(* Logix 5000 project; controller FV vendor 1 type 14 code 217 rev 31.11; software revision 31.00; part 11 of 63 *)
(* tags used below, declared in another part *)
   CWD : CHECKWORD_FLAGS;
   FR_B230 : INT[255];   // FLOW_BITS Flow Meter Bits
   FR_B240 : INT[255];   // DEBOUNCE Debounce Flags
   FR_B246 : INT[255];   // V_REVERSE Flags for reversing contol action
   FR_CFG1_P : PlantItem;   // CFG1_P
   FR_CFG2_P : PlantItem;   // CFG2_P
   FR_data_file_value_to_move : DINT;
   FR_FILT_PR_PX : PlantItem;   // FILT_PR_PX
   FR_FILT_TNK_PX : PlantItem;   // FILT_TNK_PX
   FR_FILT_TNLN_PX : PlantItem;   // FILT_TNLN_PX
   FR_FRV1_AV01 : PlantItem;   // FRV1_AV01
   FR_FV26_AV01 : PlantItem;   // FV26_AV01
   FR_FV26_AV04 : PlantItem;   // FV26_AV04
   FR_FV26_AV05 : PlantItem;   // FV26_AV05
   FR_FV26_AV06 : PlantItem;   // FV26_AV06
   FR_FV26_AV07 : PlantItem;   // FV26_AV07
   FR_FV26_VA01 : PlantItem;   // FV26_VA01
   FR_FV27_AV04 : PlantItem;   // FV27_AV04
   FR_FV28_AV04 : PlantItem;   // FV28_AV04
   FR_FV29_AV04 : PlantItem;   // FV29_AV04
   FR_FV30_AV04 : PlantItem;   // FV30_AV04
   FR_FV31_AV04 : PlantItem;   // FV31_AV04
   FR_FVR1_P01 : PlantItem;   // FVR1_P01
   FR_N10 : INT[265];   // FV_AGING Comms to FV Aging PL C
   FR_N100 : INT[265];   // FV FILLING
   FR_N110 : INT[265];   // GREEN BEER Green Beer Main
   FR_N120 : INT[265];   // YEAST CROP Yeast Cropping Main
   FR_N13 : INT[265];   // MV_ROUTE Comms to MV Routing PLC
   FR_N130 : INT[265];   // FILTRATE Filtrate Return
   FR_N14 : INT[265];   // MVFV CIP Comms to MVFV CIP Un it PLC
   FR_N160 : INT[265];   // VESSEL Vessel Working Direc tory
   FR_N200 : INT[265];   // ANALOG_IN Analog Inputs
   FR_N255 : INT[265];   // CHECKWORDS
   FR_N26 : INT[265];   // FV26
   FR_N7 : INT[265];   // INTEGER
   FR_N99 : INT[265];   // COMMENT Comment Lines
   FR_PANELESTOP : PlantItem;   // PANELESTOP
   FR_PARAF : PlantItem;   // PARAF
   FR_PILZ : PlantItem;   // PILZ
   FR_T131 : TIMER[255];   // FILTRATE
   FR_T144 : TIMER[255];   // CIP
   FR_T4 : TIMER[255];   // TIMER
   FR_VB1_AV08 : PlantItem;   // VB1_AV08
   FR_VB1_AV09 : PlantItem;   // VB1_AV09
   FR_VB4_AV01 : PlantItem;   // VB4_AV01
   FR_VB4_AV07 : PlantItem;   // VB4_AV07
   FR_VB4_AV13 : PlantItem;   // VB4_AV13
   FR_VB4_AV19 : PlantItem;   // VB4_AV19
   FR_VB4_AV21 : PlantItem;   // VB4_AV21
   FR_VB4_AV23 : PlantItem;   // VB4_AV23
(* FR_Common, continued *)

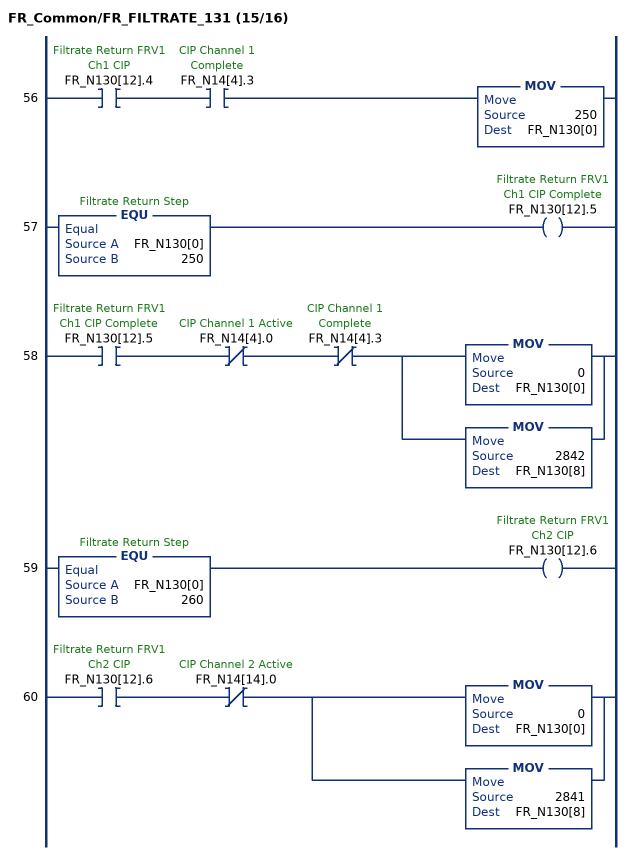
   [picture p136: FR_Common/FR_FILTRATE_131 rungs 56-60]
   56: XIC(FR_N130[12].4)XIC(FR_N14[4].3)MOV(250,FR_N130[0]);
   57: EQU(FR_N130[0],250)OTE(FR_N130[12].5);
   58: XIC(FR_N130[12].5)XIO(FR_N14[4].0)XIO(FR_N14[4].3)[MOV(0,FR_N130[0]) ,MOV(2842,FR_N130[8]) ];
   59: EQU(FR_N130[0],260)OTE(FR_N130[12].6);
   60: XIC(FR_N130[12].6)XIO(FR_N14[14].0)[MOV(0,FR_N130[0]) ,MOV(2841,FR_N130[8]) ];
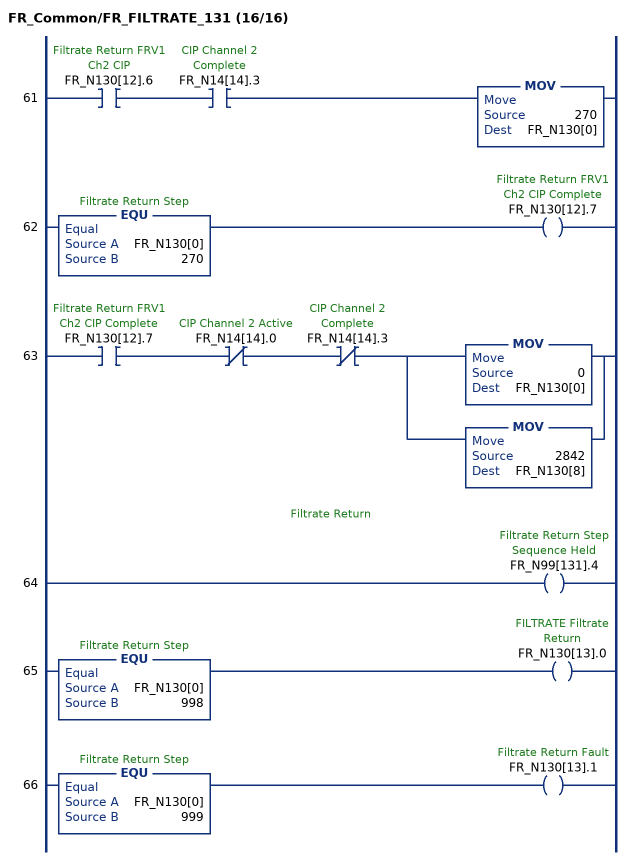
   61: XIC(FR_N130[12].6)XIC(FR_N14[14].3)MOV(270,FR_N130[0]);
   62: EQU(FR_N130[0],270)OTE(FR_N130[12].7);
   63: XIC(FR_N130[12].7)XIO(FR_N14[14].0)XIO(FR_N14[14].3)[MOV(0,FR_N130[0]) ,MOV(2842,FR_N130[8]) ];
   // Filtrate Return
   64: OTE(FR_N99[131].4);
   65: EQU(FR_N130[0],998)OTE(FR_N130[13].0);
   66: EQU(FR_N130[0],999)OTE(FR_N130[13].1);
END_ROUTINE

ROUTINE FR_FILTRATE_O_132   (* ladder *)
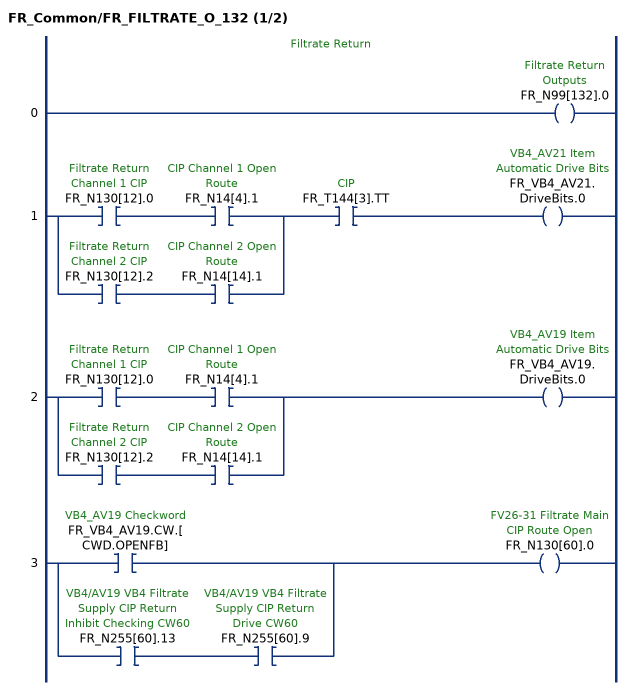
   // Filtrate Return
   0: OTE(FR_N99[132].0);
   1: [XIC(FR_N130[12].0) XIC(FR_N14[4].1) ,XIC(FR_N130[12].2) XIC(FR_N14[14].1) ]XIC(FR_T144[3].TT)OTE(FR_VB4_AV21.DriveBits.0);
   2: [XIC(FR_N130[12].0) XIC(FR_N14[4].1) ,XIC(FR_N130[12].2) XIC(FR_N14[14].1) ]OTE(FR_VB4_AV19.DriveBits.0);
   3: [XIC(FR_VB4_AV19.CW.[CWD.OPENFB]) ,XIC(FR_N255[60].13) XIC(FR_N255[60].9) ]OTE(FR_N130[60].0);
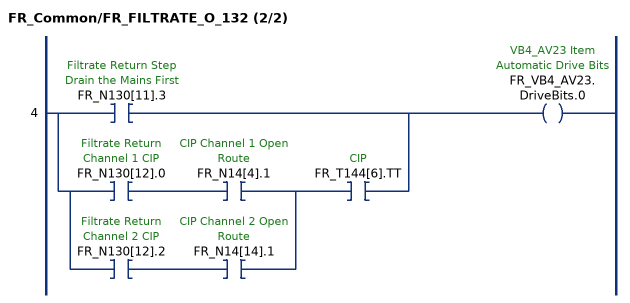
   4: [XIC(FR_N130[11].3) ,[XIC(FR_N130[12].0) XIC(FR_N14[4].1) ,XIC(FR_N130[12].2) XIC(FR_N14[14].1) ] XIC(FR_T144[6].TT) ]OTE(FR_VB4_AV23.DriveBits.0);
END_ROUTINE

ROUTINE FR_FILTRATE_S_130   (* ladder *)
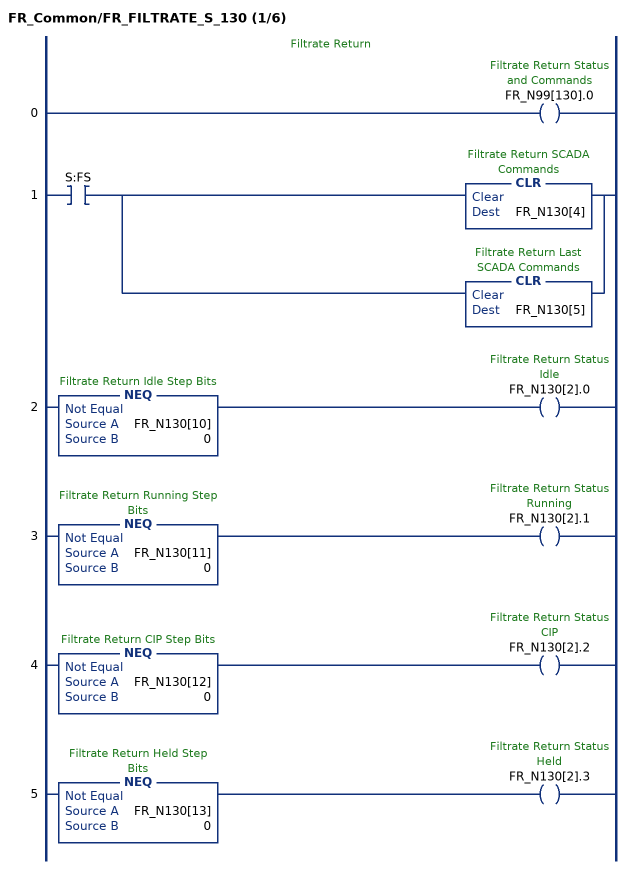
   // Filtrate Return
   0: OTE(FR_N99[130].0);
   1: XIC(S:FS)[CLR(FR_N130[4]) ,CLR(FR_N130[5]) ];
   2: NEQ(FR_N130[10],0)OTE(FR_N130[2].0);
   3: NEQ(FR_N130[11],0)OTE(FR_N130[2].1);
   4: NEQ(FR_N130[12],0)OTE(FR_N130[2].2);
   5: NEQ(FR_N130[13],0)OTE(FR_N130[2].3);
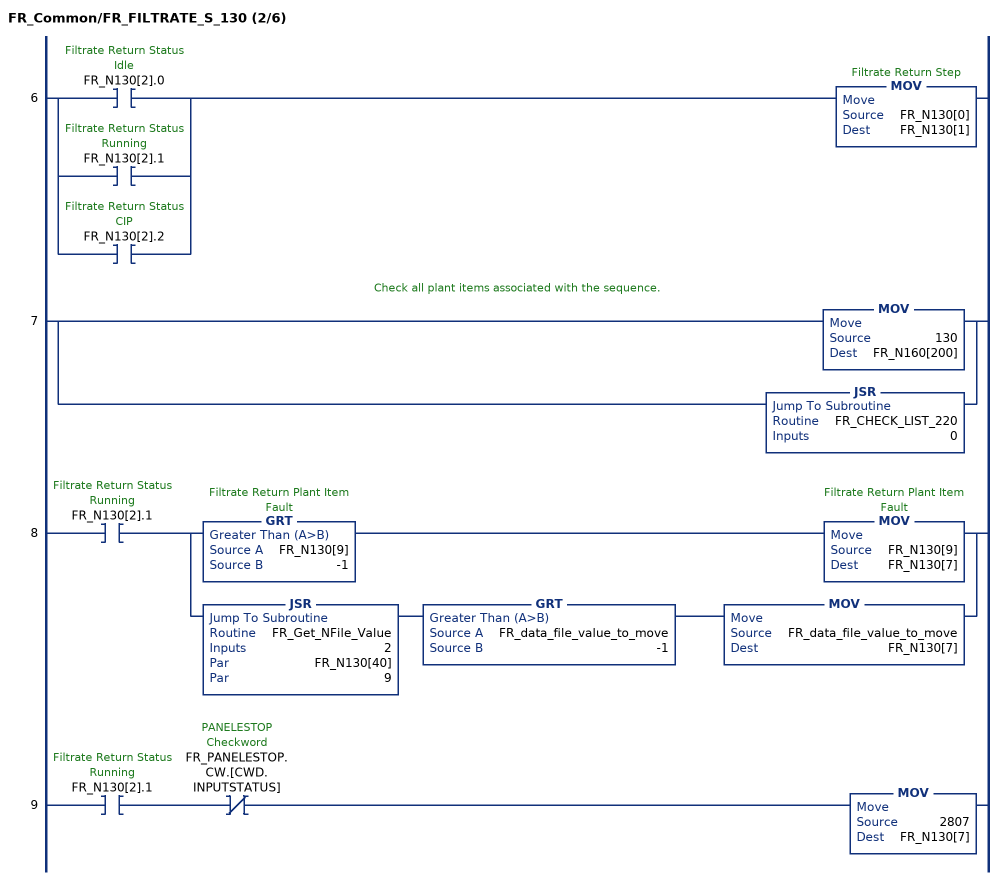
   6: [XIC(FR_N130[2].0) ,XIC(FR_N130[2].1) ,XIC(FR_N130[2].2) ]MOV(FR_N130[0],FR_N130[1]);
   // Check all plant items associated with the sequence.
   7: [MOV(130,FR_N160[200]) ,JSR(FR_CHECK_LIST_220,0) ];
   8: XIC(FR_N130[2].1)[GRT(FR_N130[9],-1) MOV(FR_N130[9],FR_N130[7]) ,JSR(FR_Get_NFile_Value,2,FR_N130[40],9) GRT(FR_data_file_value_to_move,-1) MOV(FR_data_file_value_to_move,FR_N130[7]) ];
   9: XIC(FR_N130[2].1)XIO(FR_PANELESTOP.CW.[CWD.INPUTSTATUS])MOV(2807,FR_N130[7]);
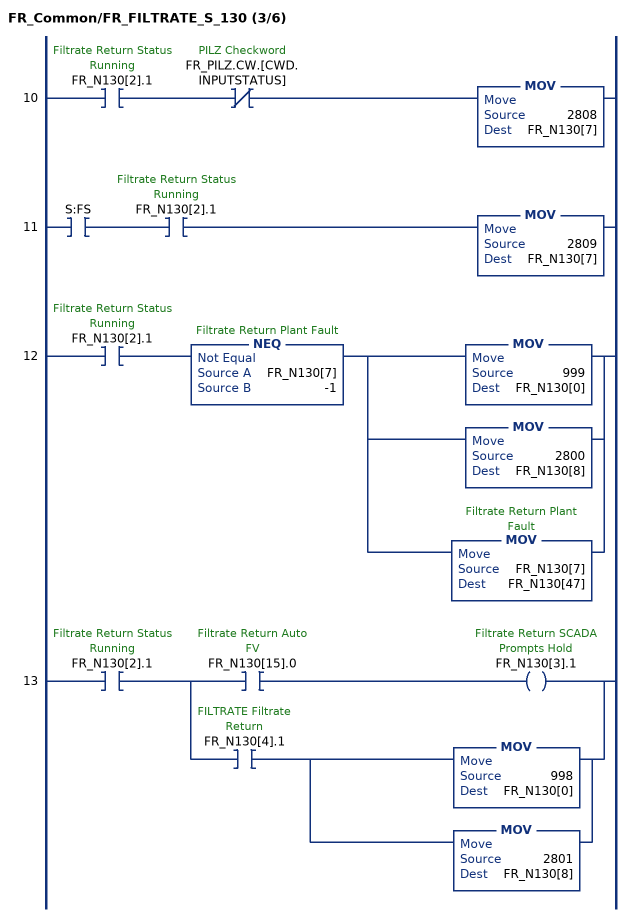
   10: XIC(FR_N130[2].1)XIO(FR_PILZ.CW.[CWD.INPUTSTATUS])MOV(2808,FR_N130[7]);
   11: XIC(S:FS)XIC(FR_N130[2].1)MOV(2809,FR_N130[7]);
   12: XIC(FR_N130[2].1)NEQ(FR_N130[7],-1)[MOV(999,FR_N130[0]) ,MOV(2800,FR_N130[8]) ,MOV(FR_N130[7],FR_N130[47]) ];
   13: XIC(FR_N130[2].1)[XIC(FR_N130[15].0) OTE(FR_N130[3].1) ,XIC(FR_N130[4].1) [MOV(998,FR_N130[0]) ,MOV(2801,FR_N130[8]) ] ];
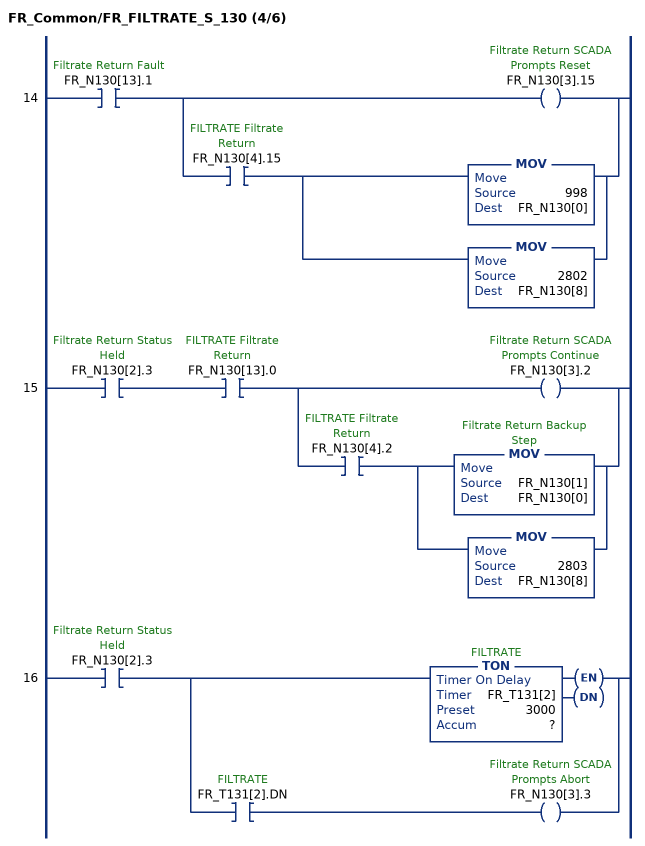
   14: XIC(FR_N130[13].1)[OTE(FR_N130[3].15) ,XIC(FR_N130[4].15) [MOV(998,FR_N130[0]) ,MOV(2802,FR_N130[8]) ] ];
   15: XIC(FR_N130[2].3)XIC(FR_N130[13].0)[OTE(FR_N130[3].2) ,XIC(FR_N130[4].2) [MOV(FR_N130[1],FR_N130[0]) ,MOV(2803,FR_N130[8]) ] ];
   16: XIC(FR_N130[2].3)[TON(FR_T131[2],?,?) ,XIC(FR_T131[2].DN) OTE(FR_N130[3].3) ];
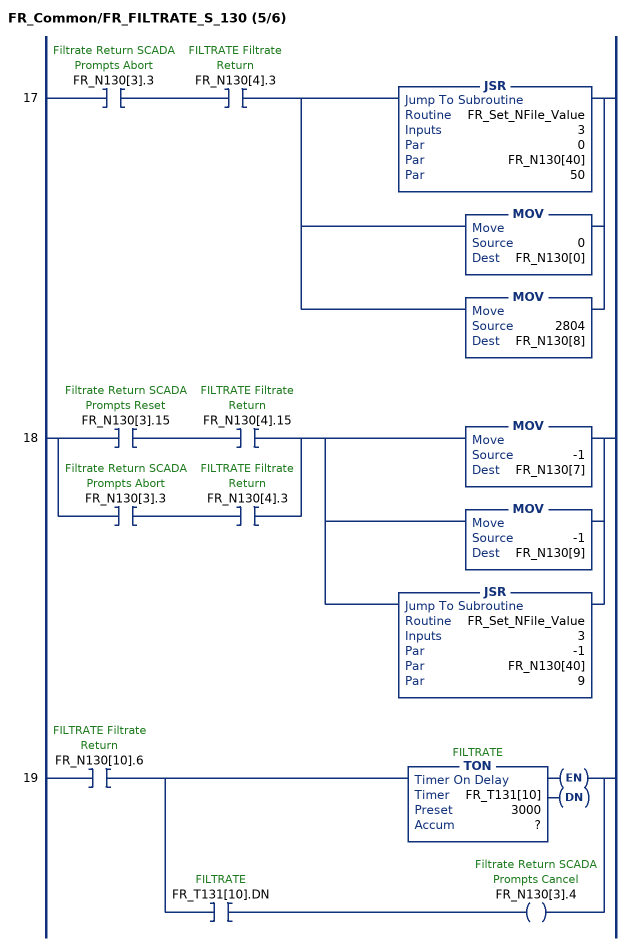
   17: XIC(FR_N130[3].3)XIC(FR_N130[4].3)[JSR(FR_Set_NFile_Value,3,0,FR_N130[40],50) ,MOV(0,FR_N130[0]) ,MOV(2804,FR_N130[8]) ];
   18: [XIC(FR_N130[3].15) XIC(FR_N130[4].15) ,XIC(FR_N130[3].3) XIC(FR_N130[4].3) ][MOV(-1,FR_N130[7]) ,MOV(-1,FR_N130[9]) ,JSR(FR_Set_NFile_Value,3,-1,FR_N130[40],9) ];
   19: XIC(FR_N130[10].6)[TON(FR_T131[10],?,?) ,XIC(FR_T131[10].DN) OTE(FR_N130[3].4) ];
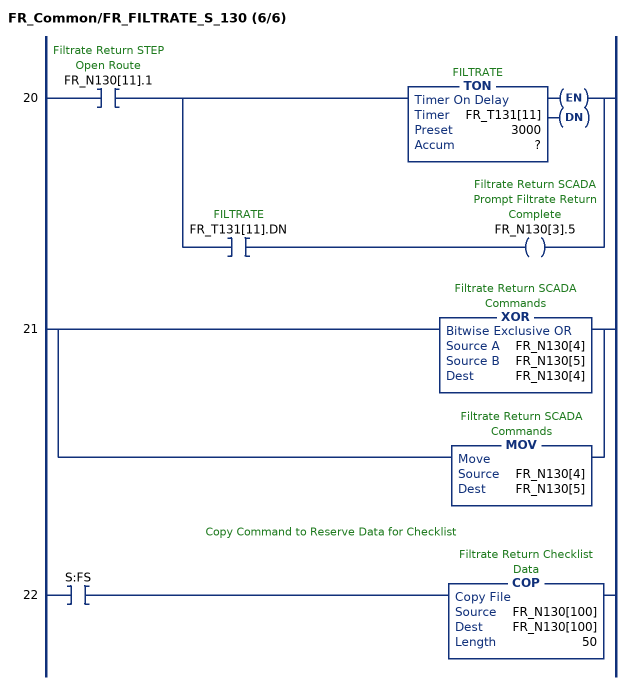
   20: XIC(FR_N130[11].1)[TON(FR_T131[11],?,?) ,XIC(FR_T131[11].DN) OTE(FR_N130[3].5) ];
   21: [XOR(FR_N130[4],FR_N130[5],FR_N130[4]) ,MOV(FR_N130[4],FR_N130[5]) ];
   // Copy Command to Reserve Data for Checklist
   22: XIC(S:FS)COP(FR_N130[100],FR_N130[100],50);
END_ROUTINE

ROUTINE FR_FLOWMETER_230   (* ladder *)
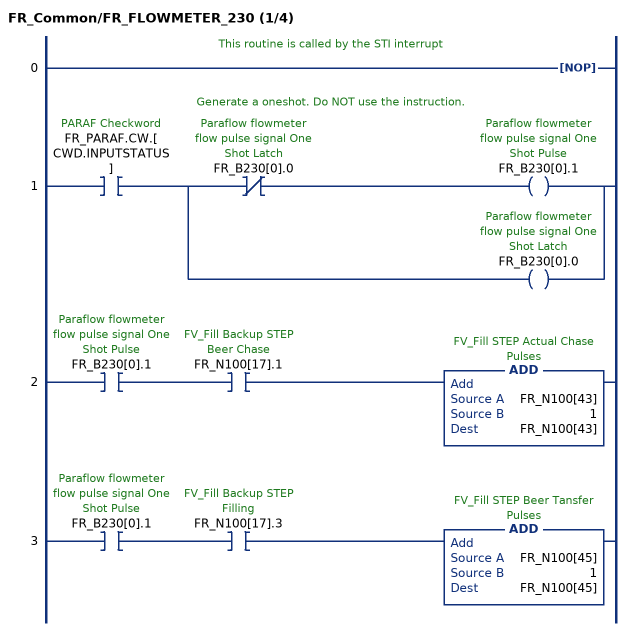
   // This routine is called by the STI interrupt
   0: NOP();
   // Generate a oneshot. Do NOT use the instruction.
   1: XIC(FR_PARAF.CW.[CWD.INPUTSTATUS])[XIO(FR_B230[0].0) OTE(FR_B230[0].1) ,OTE(FR_B230[0].0) ];
   2: XIC(FR_B230[0].1)XIC(FR_N100[17].1)ADD(FR_N100[43],1,FR_N100[43]);
   3: XIC(FR_B230[0].1)XIC(FR_N100[17].3)ADD(FR_N100[45],1,FR_N100[45]);
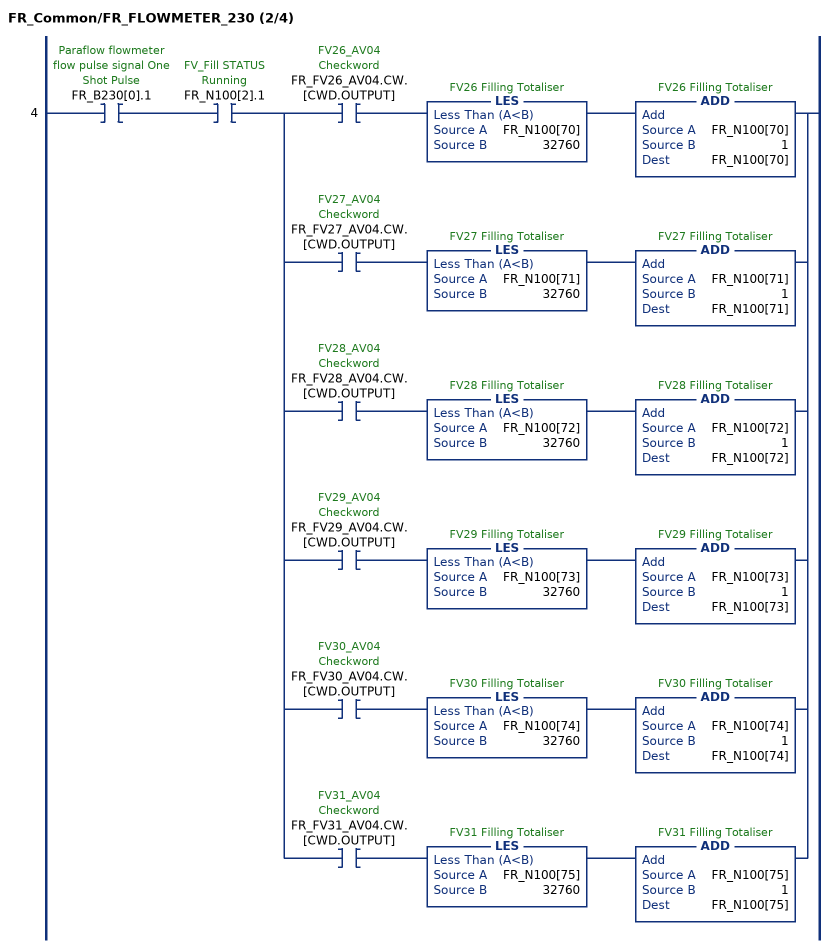
   4: XIC(FR_B230[0].1)XIC(FR_N100[2].1)[XIC(FR_FV26_AV04.CW.[CWD.OUTPUT]) LES(FR_N100[70],32760) ADD(FR_N100[70],1,FR_N100[70]) ,XIC(FR_FV27_AV04.CW.[CWD.OUTPUT]) LES(FR_N100[71],32760) ADD(FR_N100[71],1,FR_N100[71]) ,XIC(FR_FV28_AV04.CW.[CWD.OUTPUT]) LES(FR_N100[72],32760) ADD(FR_N100[72],1,FR_N100[72]) ,XIC(FR_FV29_AV04.CW.[CWD.OUTPUT]) LES(FR_N100[73],32760) ADD(FR_N100[73],1,FR_N100[73]) ,XIC(FR_FV30_AV04.CW.[CWD.OUTPUT]) LES(FR_N100[74],32760) ADD(FR_N100[74],1,FR_N100[74]) ,XIC(FR_FV31_AV04.CW.[CWD.OUTPUT]) LES(FR_N100[75],32760) ADD(FR_N100[75],1,FR_N100[75]) ];
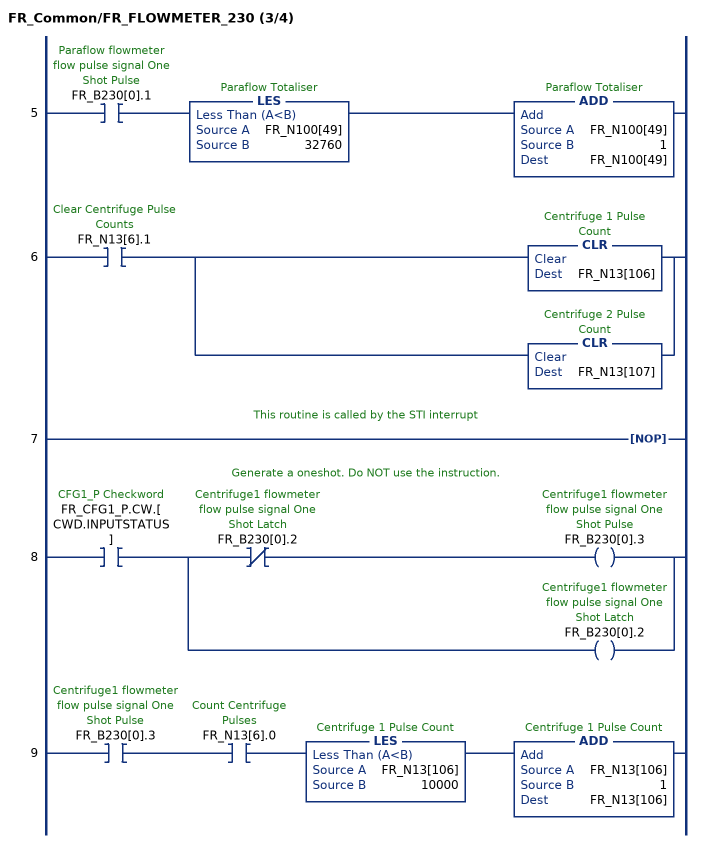
   5: XIC(FR_B230[0].1)LES(FR_N100[49],32760)ADD(FR_N100[49],1,FR_N100[49]);
   6: XIC(FR_N13[6].1)[CLR(FR_N13[106]) ,CLR(FR_N13[107]) ];
   // This routine is called by the STI interrupt
   7: NOP();
   // Generate a oneshot. Do NOT use the instruction.
   8: XIC(FR_CFG1_P.CW.[CWD.INPUTSTATUS])[XIO(FR_B230[0].2) OTE(FR_B230[0].3) ,OTE(FR_B230[0].2) ];
   9: XIC(FR_B230[0].3)XIC(FR_N13[6].0)LES(FR_N13[106],10000)ADD(FR_N13[106],1,FR_N13[106]);
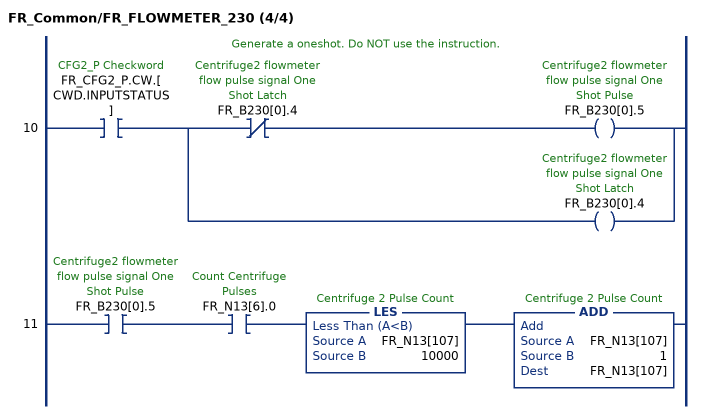
   // Generate a oneshot. Do NOT use the instruction.
   10: XIC(FR_CFG2_P.CW.[CWD.INPUTSTATUS])[XIO(FR_B230[0].4) OTE(FR_B230[0].5) ,OTE(FR_B230[0].4) ];
   11: XIC(FR_B230[0].5)XIC(FR_N13[6].0)LES(FR_N13[107],10000)ADD(FR_N13[107],1,FR_N13[107]);
END_ROUTINE

ROUTINE FR_FRV_133   (* ladder *)
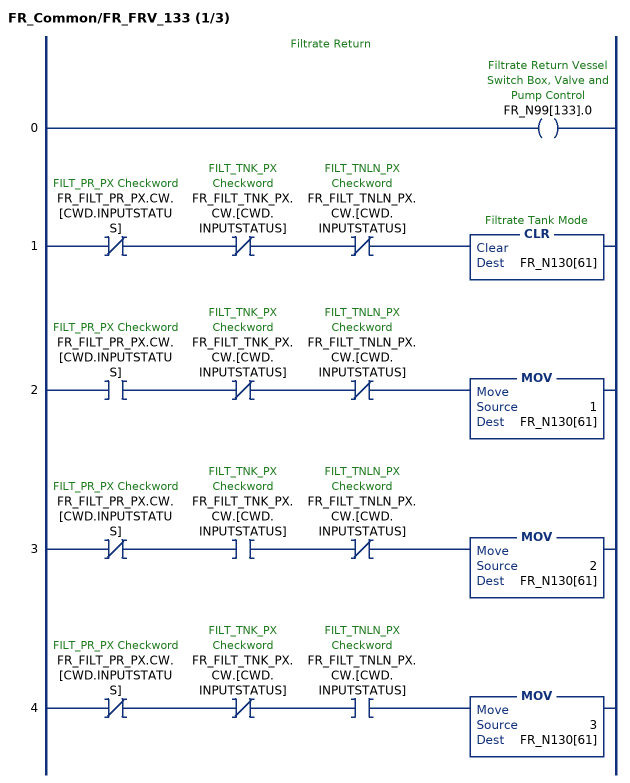
   // Filtrate Return
   0: OTE(FR_N99[133].0);
   1: XIO(FR_FILT_PR_PX.CW.[CWD.INPUTSTATUS])XIO(FR_FILT_TNK_PX.CW.[CWD.INPUTSTATUS])XIO(FR_FILT_TNLN_PX.CW.[CWD.INPUTSTATUS])CLR(FR_N130[61]);
   2: XIC(FR_FILT_PR_PX.CW.[CWD.INPUTSTATUS])XIO(FR_FILT_TNK_PX.CW.[CWD.INPUTSTATUS])XIO(FR_FILT_TNLN_PX.CW.[CWD.INPUTSTATUS])MOV(1,FR_N130[61]);
   3: XIO(FR_FILT_PR_PX.CW.[CWD.INPUTSTATUS])XIC(FR_FILT_TNK_PX.CW.[CWD.INPUTSTATUS])XIO(FR_FILT_TNLN_PX.CW.[CWD.INPUTSTATUS])MOV(2,FR_N130[61]);
   4: XIO(FR_FILT_PR_PX.CW.[CWD.INPUTSTATUS])XIO(FR_FILT_TNK_PX.CW.[CWD.INPUTSTATUS])XIC(FR_FILT_TNLN_PX.CW.[CWD.INPUTSTATUS])MOV(3,FR_N130[61]);
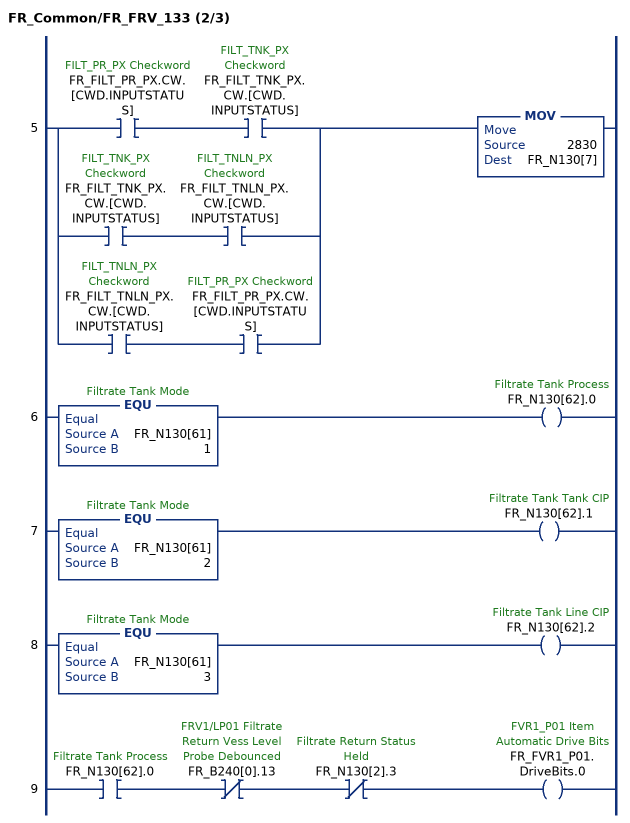
   5: [XIC(FR_FILT_PR_PX.CW.[CWD.INPUTSTATUS]) XIC(FR_FILT_TNK_PX.CW.[CWD.INPUTSTATUS]) ,XIC(FR_FILT_TNK_PX.CW.[CWD.INPUTSTATUS]) XIC(FR_FILT_TNLN_PX.CW.[CWD.INPUTSTATUS]) ,XIC(FR_FILT_TNLN_PX.CW.[CWD.INPUTSTATUS]) XIC(FR_FILT_PR_PX.CW.[CWD.INPUTSTATUS]) ]MOV(2830,FR_N130[7]);
   6: EQU(FR_N130[61],1)OTE(FR_N130[62].0);
   7: EQU(FR_N130[61],2)OTE(FR_N130[62].1);
   8: EQU(FR_N130[61],3)OTE(FR_N130[62].2);
   9: XIC(FR_N130[62].0)XIO(FR_B240[0].13)XIO(FR_N130[2].3)OTE(FR_FVR1_P01.DriveBits.0);
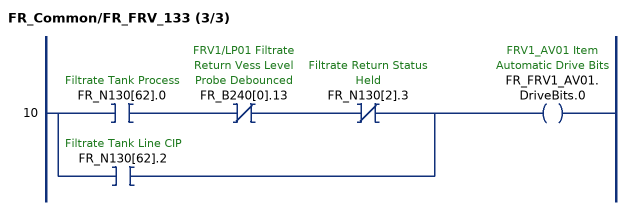
   10: [XIC(FR_N130[62].0) XIO(FR_B240[0].13) XIO(FR_N130[2].3) ,XIC(FR_N130[62].2) ]OTE(FR_FRV1_AV01.DriveBits.0);
END_ROUTINE

ROUTINE FR_FV26_26   (* ladder *)
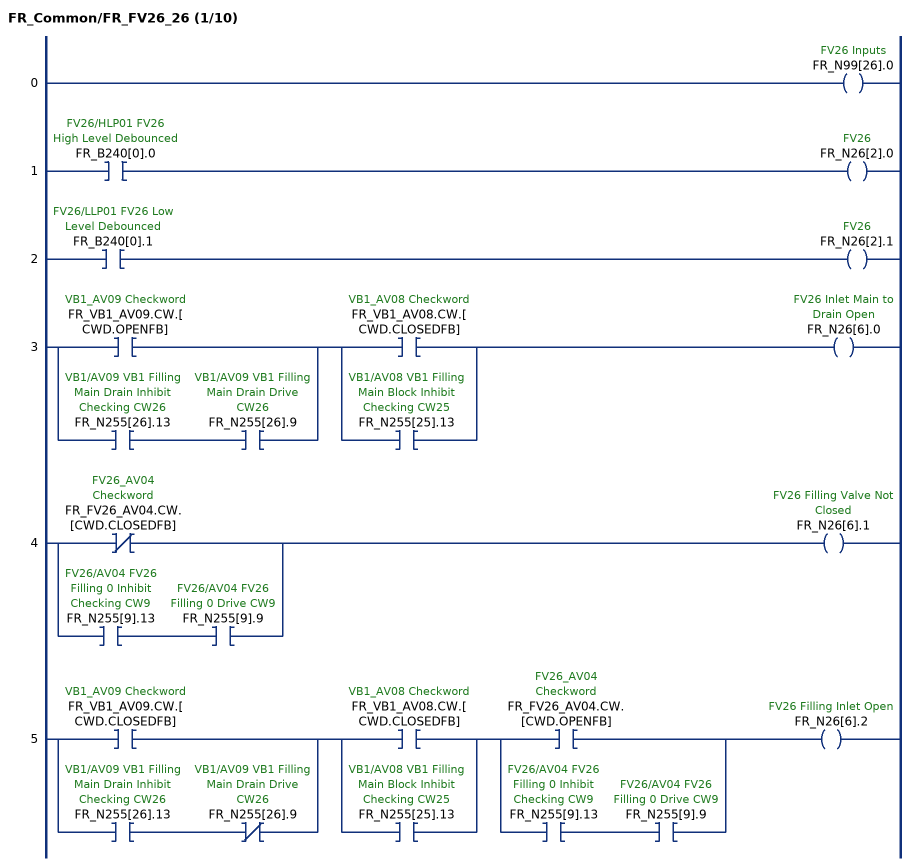
   0: OTE(FR_N99[26].0);
   1: XIC(FR_B240[0].0)OTE(FR_N26[2].0);
   2: XIC(FR_B240[0].1)OTE(FR_N26[2].1);
   3: [XIC(FR_VB1_AV09.CW.[CWD.OPENFB]) ,XIC(FR_N255[26].13) XIC(FR_N255[26].9) ][XIC(FR_VB1_AV08.CW.[CWD.CLOSEDFB]) ,XIC(FR_N255[25].13) ]OTE(FR_N26[6].0);
   4: [XIO(FR_FV26_AV04.CW.[CWD.CLOSEDFB]) ,XIC(FR_N255[9].13) XIC(FR_N255[9].9) ]OTE(FR_N26[6].1);
   5: [XIC(FR_VB1_AV09.CW.[CWD.CLOSEDFB]) ,XIC(FR_N255[26].13) XIO(FR_N255[26].9) ][XIC(FR_VB1_AV08.CW.[CWD.CLOSEDFB]) ,XIC(FR_N255[25].13) ][XIC(FR_FV26_AV04.CW.[CWD.OPENFB]) ,XIC(FR_N255[9].13) XIC(FR_N255[9].9) ]OTE(FR_N26[6].2);
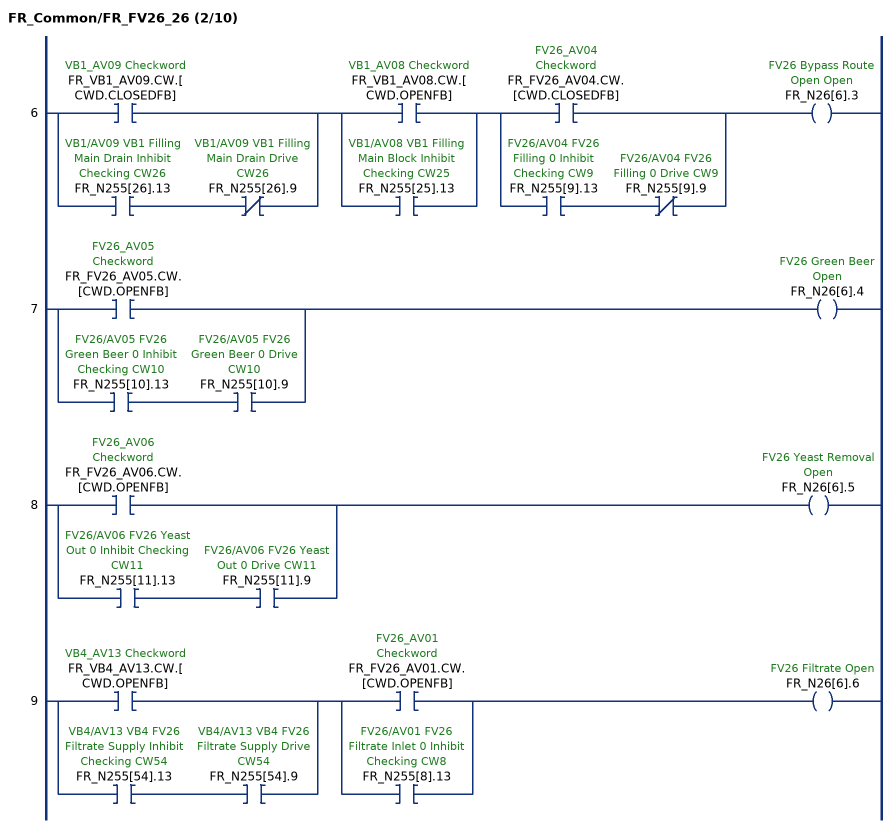
   6: [XIC(FR_VB1_AV09.CW.[CWD.CLOSEDFB]) ,XIC(FR_N255[26].13) XIO(FR_N255[26].9) ][XIC(FR_VB1_AV08.CW.[CWD.OPENFB]) ,XIC(FR_N255[25].13) ][XIC(FR_FV26_AV04.CW.[CWD.CLOSEDFB]) ,XIC(FR_N255[9].13) XIO(FR_N255[9].9) ]OTE(FR_N26[6].3);
   7: [XIC(FR_FV26_AV05.CW.[CWD.OPENFB]) ,XIC(FR_N255[10].13) XIC(FR_N255[10].9) ]OTE(FR_N26[6].4);
   8: [XIC(FR_FV26_AV06.CW.[CWD.OPENFB]) ,XIC(FR_N255[11].13) XIC(FR_N255[11].9) ]OTE(FR_N26[6].5);
   9: [XIC(FR_VB4_AV13.CW.[CWD.OPENFB]) ,XIC(FR_N255[54].13) XIC(FR_N255[54].9) ][XIC(FR_FV26_AV01.CW.[CWD.OPENFB]) ,XIC(FR_N255[8].13) ]OTE(FR_N26[6].6);
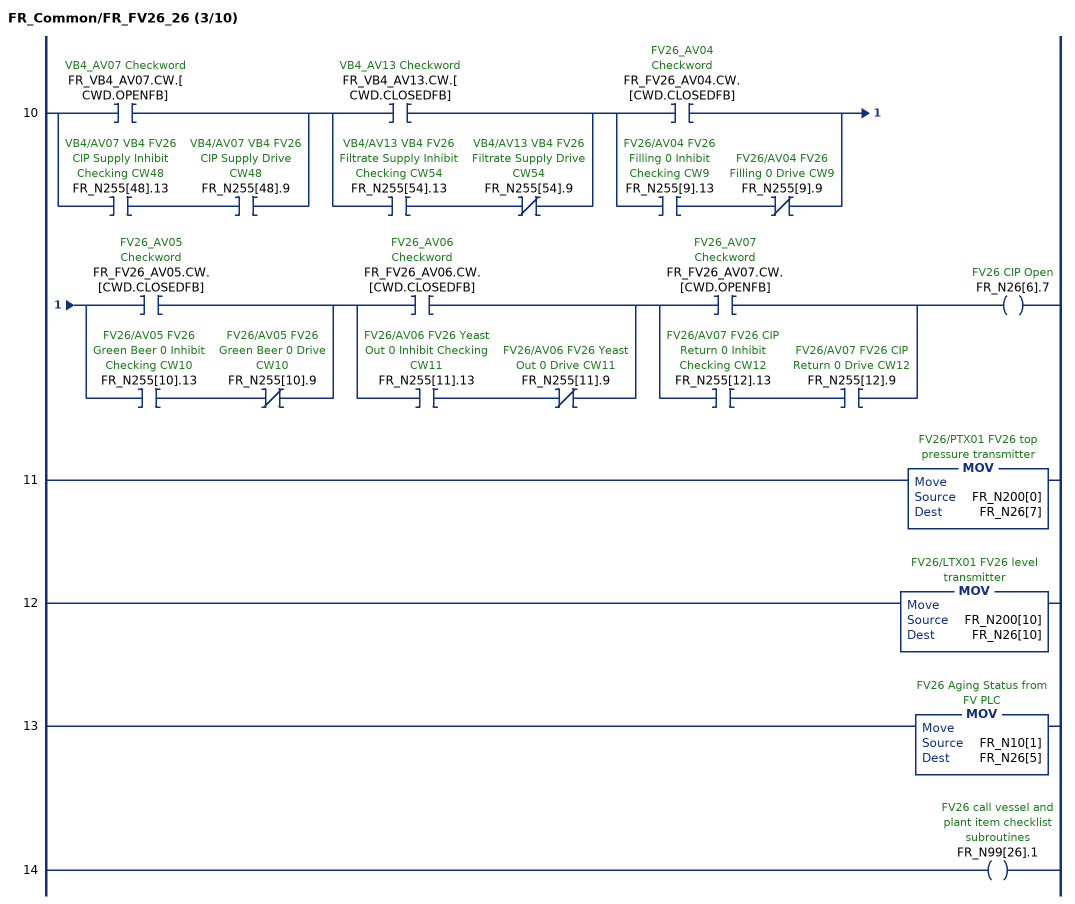
   10: [XIC(FR_VB4_AV07.CW.[CWD.OPENFB]) ,XIC(FR_N255[48].13) XIC(FR_N255[48].9) ][XIC(FR_VB4_AV13.CW.[CWD.CLOSEDFB]) ,XIC(FR_N255[54].13) XIO(FR_N255[54].9) ][XIC(FR_FV26_AV04.CW.[CWD.CLOSEDFB]) ,XIC(FR_N255[9].13) XIO(FR_N255[9].9) ][XIC(FR_FV26_AV05.CW.[CWD.CLOSEDFB]) ,XIC(FR_N255[10].13) XIO(FR_N255[10].9) ][XIC(FR_FV26_AV06.CW.[CWD.CLOSEDFB]) ,XIC(FR_N255[11].13) XIO(FR_N255[11].9) ][XIC(FR_FV26_AV07.CW.[CWD.OPENFB]) ,XIC(FR_N255[12].13) XIC(FR_N255[12].9) ]OTE(FR_N26[6].7);
   11: MOV(FR_N200[0],FR_N26[7]);
   12: MOV(FR_N200[10],FR_N26[10]);
   13: MOV(FR_N10[1],FR_N26[5]);
   14: OTE(FR_N99[26].1);
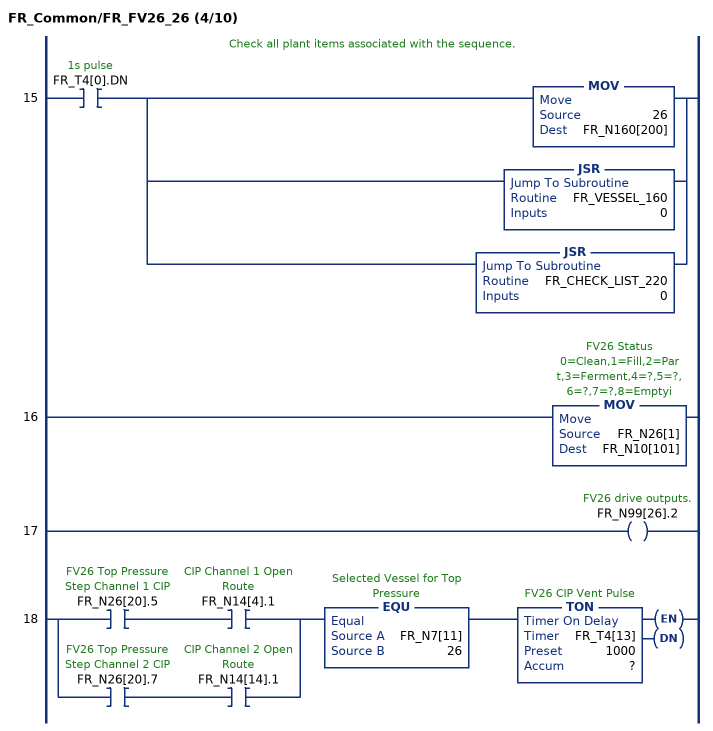
   // Check all plant items associated with the sequence.
   15: XIC(FR_T4[0].DN)[MOV(26,FR_N160[200]) ,JSR(FR_VESSEL_160,0) ,JSR(FR_CHECK_LIST_220,0) ];
   16: MOV(FR_N26[1],FR_N10[101]);
   17: OTE(FR_N99[26].2);
   18: [XIC(FR_N26[20].5) XIC(FR_N14[4].1) ,XIC(FR_N26[20].7) XIC(FR_N14[14].1) ]EQU(FR_N7[11],26)TON(FR_T4[13],?,?);
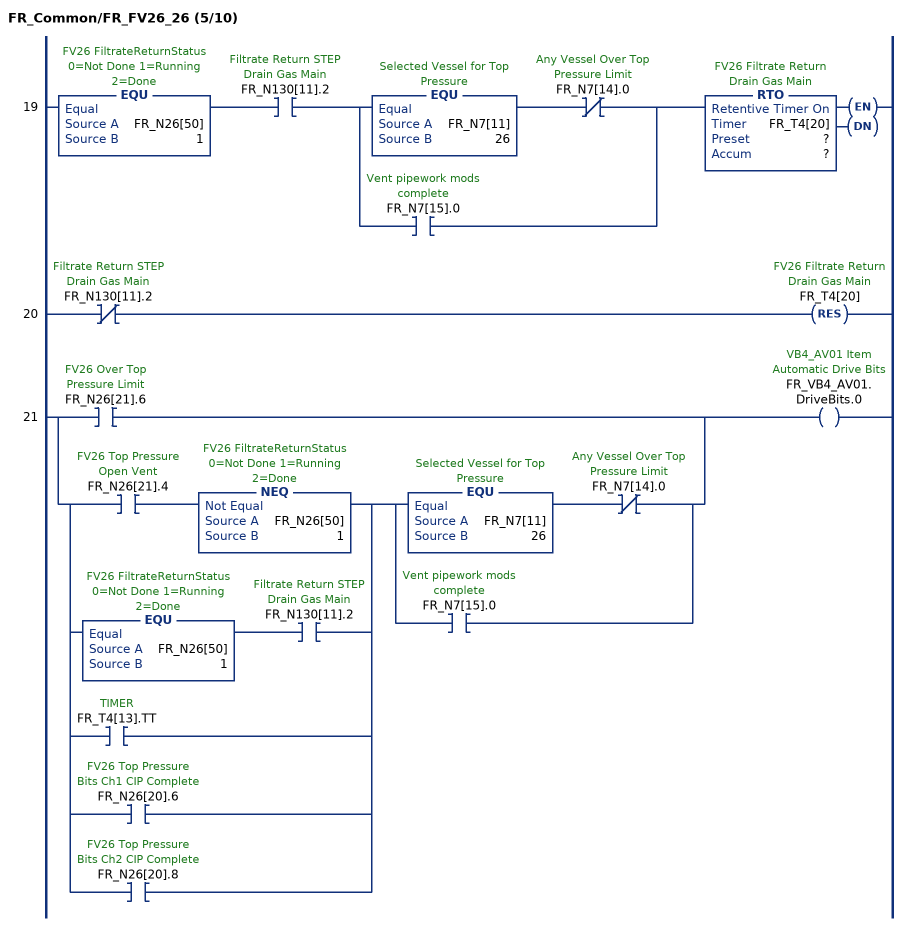
   19: EQU(FR_N26[50],1)XIC(FR_N130[11].2)[EQU(FR_N7[11],26) XIO(FR_N7[14].0) ,XIC(FR_N7[15].0) ]RTO(FR_T4[20],?,?);
   20: XIO(FR_N130[11].2)RES(FR_T4[20]);
   21: [XIC(FR_N26[21].6) ,[XIC(FR_N26[21].4) NEQ(FR_N26[50],1) ,EQU(FR_N26[50],1) XIC(FR_N130[11].2) ,XIC(FR_T4[13].TT) ,[XIC(FR_N26[20].6) ,XIC(FR_N26[20].8) ] ] [EQU(FR_N7[11],26) XIO(FR_N7[14].0) ,XIC(FR_N7[15].0) ] ]OTE(FR_VB4_AV01.DriveBits.0);
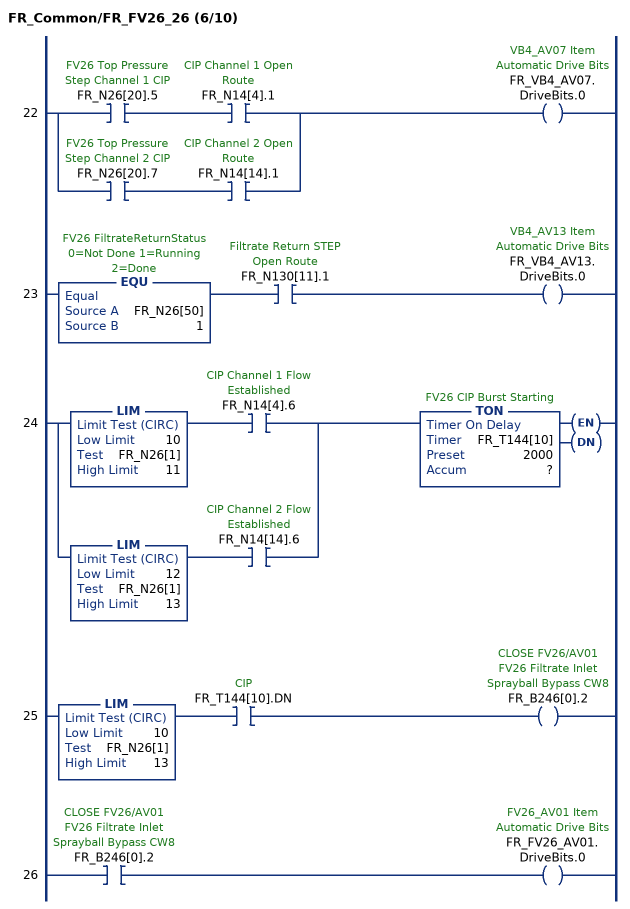
   22: [XIC(FR_N26[20].5) XIC(FR_N14[4].1) ,XIC(FR_N26[20].7) XIC(FR_N14[14].1) ]OTE(FR_VB4_AV07.DriveBits.0);
   23: EQU(FR_N26[50],1)XIC(FR_N130[11].1)OTE(FR_VB4_AV13.DriveBits.0);
   24: [LIM(10,FR_N26[1],11) XIC(FR_N14[4].6) ,LIM(12,FR_N26[1],13) XIC(FR_N14[14].6) ]TON(FR_T144[10],?,?);
   25: LIM(10,FR_N26[1],13)XIC(FR_T144[10].DN)OTE(FR_B246[0].2);
   26: XIC(FR_B246[0].2)OTE(FR_FV26_AV01.DriveBits.0);
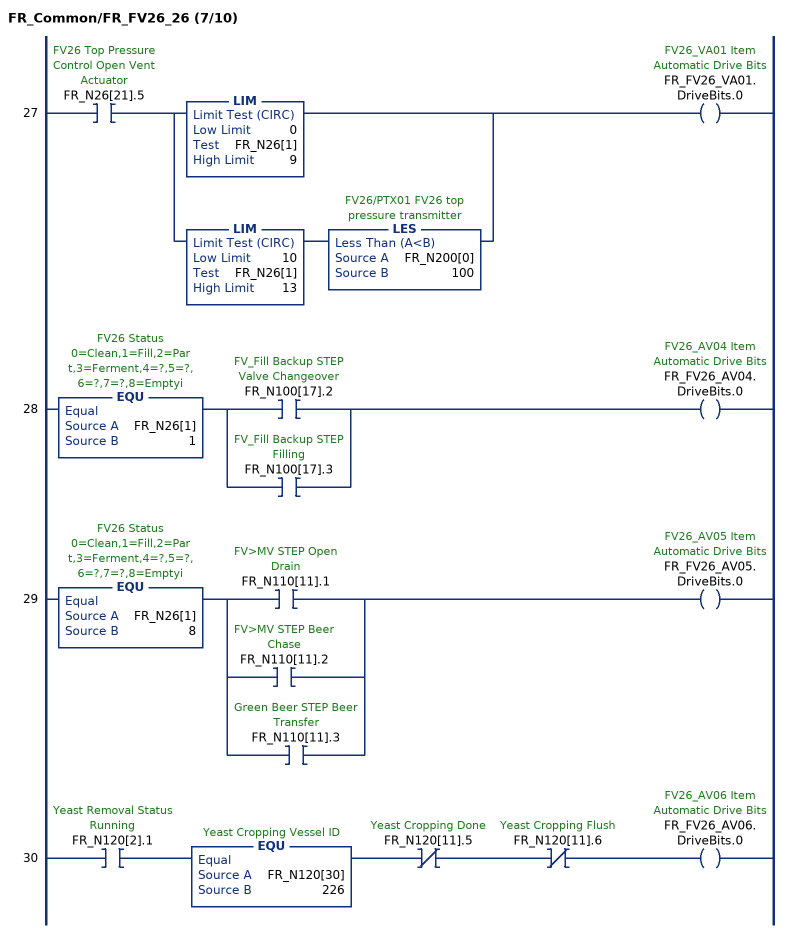
   27: XIC(FR_N26[21].5)[LIM(0,FR_N26[1],9) ,LIM(10,FR_N26[1],13) LES(FR_N200[0],100) ]OTE(FR_FV26_VA01.DriveBits.0);
   28: EQU(FR_N26[1],1)[XIC(FR_N100[17].2) ,XIC(FR_N100[17].3) ]OTE(FR_FV26_AV04.DriveBits.0);
   29: EQU(FR_N26[1],8)[XIC(FR_N110[11].1) ,XIC(FR_N110[11].2) ,XIC(FR_N110[11].3) ]OTE(FR_FV26_AV05.DriveBits.0);
   30: XIC(FR_N120[2].1)EQU(FR_N120[30],226)XIO(FR_N120[11].5)XIO(FR_N120[11].6)OTE(FR_FV26_AV06.DriveBits.0);
